(* Logix 5000 project; controller PLC_MCC1300_75F1 vendor 1 type 14 code 166 rev 32.11; software revision 32.04; part 40 of 83 *)
(* tags used below, declared in another part *)
   CONST_rgdDestMask : DINT[32];   // Destination Mask
   GP_RampSpace : GP_RampSpace;
   I : INT[128];   // Local Input Updates Input Slot 2
   TMP_d : DINT;
   TMP_dConv : DINT;
   TMP_dEndConveyorPos : DINT;
   TMP_dIndexMotor : DINT;
   TMP_dIndexNext : DINT;
   TMP_dIndexPrevious : DINT;
   TMP_dTailOnNextConveyor_cmm : DINT;
   TMP_xLastConv : BOOL;
   TMP_xOSN : DINT;
   TMP_xOSN_B : DINT;
   TMP_xOSR : DINT;
   TMP_xOSR_B : DINT;
   TMP_xSimulationActive : BOOL;
   xAlwaysOFF : BOOL;
   xAlwaysON : BOOL;
   xDebugOFF : BOOL;
   xDebugON : BOOL;
   Z300_Conveyor : UDT_StandConv[29];
   Z300_Conveyor_ALM : MAC_Conveyor_ZC_ALM[29];
   Z300_Conveyor_Conf : UDT_Conveyor_Config[29];
   Z300_Conveyor_HMW : MAC_Conveyor_ZC_HMW[29];
   Z300_Conveyor_IN_MOTION : MAC_Conveyor_ZC_IN_MOTION[29];
   Z300_LineTracking : UDT_LINE_TRACKING;
   Z301 : MAC_Zone_ML;
(* MainProgram, continued *)

ROUTINE Conv_Config   (* structured text *)
   //// CONVEYORS CONFIGURATION ////
   
   //M2CM01 (M302M1)
   Z300_Conveyor_Conf[0].dLengthConveyor_cmm := 45000;
   Z300_Conveyor_Conf[0].dWidthConveyor_cmm := 450000;
   Z300_Conveyor_Conf[0].dPitchRoller := 25000;
   Z300_Conveyor_Conf[0].dSpaceRestartPlate_cmm := 0;
   Z300_Conveyor_Conf[0].dMachineIndex := 0;
   Z300_Conveyor_Conf[0].dZoneConveyor := 1; //Z301
   Z300_Conveyor_Conf[0].dMotorNumber := 0; //Single motor
   Z300_Conveyor_Conf[0].dIndexMainSpeed := 1; //Lehr speed
   Z300_Conveyor_Conf[0].xContinuousConveyor := 1;
   Z300_Conveyor_Conf[0].xWaitGlassForStop := 0;
   Z300_Conveyor_Conf[0].rAccH_ms2 := 1.2;
   Z300_Conveyor_Conf[0].rDecH_ms2 := 1.2;
   Z300_Conveyor_Conf[0].rAccH_s := 0.75; //acceleration time with max speed 54 m/min
   Z300_Conveyor_Conf[0].rDecH_s := 0.75; //acceleration time with max speed 54 m/min
   Z300_Conveyor_Conf[0].rAccL_ms2 := 0.7;
   Z300_Conveyor_Conf[0].rDecL_ms2 := 0.7;
   Z300_Conveyor_Conf[0].rAccL_s := 1.29; //acceleration time with max speed 54 m/min
   Z300_Conveyor_Conf[0].rDecL_s := 1.29; //acceleration time with max speed 54 m/min
   Z300_Conveyor_Conf[0].xSimulationMotor := TMP_xSimulationActive;
   Z300_Conveyor_Conf[0].xLocalCleaningAllow := 0;
   Z300_Conveyor_Conf[0].xOnlyOnePlateAtTheTime := 0;
   Z300_Conveyor_Conf[0].rgxAllowedDest := CONST_rgdDestMask[0] AND CONST_rgdDestMask[1] AND CONST_rgdDestMask[2] AND CONST_rgdDestMask[3] AND CONST_rgdDestMask[4] AND CONST_rgdDestMask[5] AND CONST_rgdDestMask[6];
   Z300_Conveyor_Conf[0].rgxAllowedCullet := CONST_rgdDestMask[24];
   Z300_Conveyor_Conf[0].rgxAllowedQuality := CONST_rgdDestMask[29] AND CONST_rgdDestMask[30] AND CONST_rgdDestMask[31];
   Z300_Conveyor[0].tmOFF_DriveEnable[0].PRE := 30000;
   Z300_Conveyor[0].tmON_FeedbackTimeout[0].PRE := 2500;
   Z300_Conveyor[0].tmON_DelayReadyToMove[0].PRE := 200;
   Z300_Conveyor[0].tmON_FeedbackDriveReady[0].PRE := 1000;
   
   //M2CM02 (M302M2)
   Z300_Conveyor_Conf[1].dLengthConveyor_cmm := 31000;
   Z300_Conveyor_Conf[1].dWidthConveyor_cmm := 450000;
   Z300_Conveyor_Conf[1].dPitchRoller := 25000;
   Z300_Conveyor_Conf[1].dSpaceRestartPlate_cmm := 0;
   Z300_Conveyor_Conf[1].dMachineIndex := 1;
   Z300_Conveyor_Conf[1].dZoneConveyor := 1; //Z301
   Z300_Conveyor_Conf[1].dMotorNumber := 0; //Single motor
   Z300_Conveyor_Conf[1].dIndexMainSpeed := 1; //Lehr speed
   Z300_Conveyor_Conf[1].xContinuousConveyor := 1;
   Z300_Conveyor_Conf[1].xWaitGlassForStop := 0;
   Z300_Conveyor_Conf[1].rAccH_ms2 := 1.2;
   Z300_Conveyor_Conf[1].rDecH_ms2 := 1.2;
   Z300_Conveyor_Conf[1].rAccH_s := 0.75; //acceleration time with max speed 54 m/min
   Z300_Conveyor_Conf[1].rDecH_s := 0.75; //acceleration time with max speed 54 m/min
   Z300_Conveyor_Conf[1].rAccL_ms2 := 0.7;
   Z300_Conveyor_Conf[1].rDecL_ms2 := 0.7;
   Z300_Conveyor_Conf[1].rAccL_s := 1.29; //acceleration time with max speed 54 m/min
   Z300_Conveyor_Conf[1].rDecL_s := 1.29; //acceleration time with max speed 54 m/min
   Z300_Conveyor_Conf[1].xSimulationMotor := TMP_xSimulationActive;
   Z300_Conveyor_Conf[1].xLocalCleaningAllow := 0;
   Z300_Conveyor_Conf[1].xOnlyOnePlateAtTheTime := 0;
   Z300_Conveyor_Conf[1].rgxAllowedDest := CONST_rgdDestMask[0] AND CONST_rgdDestMask[1] AND CONST_rgdDestMask[2] AND CONST_rgdDestMask[3] AND CONST_rgdDestMask[4] AND CONST_rgdDestMask[5] AND CONST_rgdDestMask[6];
   Z300_Conveyor_Conf[1].rgxAllowedCullet := CONST_rgdDestMask[24];
   Z300_Conveyor_Conf[1].rgxAllowedQuality := CONST_rgdDestMask[29] AND CONST_rgdDestMask[30] AND CONST_rgdDestMask[31];
   Z300_Conveyor[1].tmOFF_DriveEnable[0].PRE := 30000;
   Z300_Conveyor[1].tmON_FeedbackTimeout[0].PRE := 2500;
   Z300_Conveyor[1].tmON_DelayReadyToMove[0].PRE := 200;
   Z300_Conveyor[1].tmON_FeedbackDriveReady[0].PRE := 1000;
   
   //M2CM03 (M302M3)
   Z300_Conveyor_Conf[2].dLengthConveyor_cmm := 16000;
   Z300_Conveyor_Conf[2].dWidthConveyor_cmm := 450000;
   Z300_Conveyor_Conf[2].dPitchRoller := 25000;
   Z300_Conveyor_Conf[2].dSpaceRestartPlate_cmm := 0;
   Z300_Conveyor_Conf[2].dMachineIndex := 2;
   Z300_Conveyor_Conf[2].dZoneConveyor := 1; //Z301
   Z300_Conveyor_Conf[2].dMotorNumber := 0; //Single motor
   Z300_Conveyor_Conf[2].dIndexMainSpeed := 1; //Lehr speed
   Z300_Conveyor_Conf[2].xContinuousConveyor := 1;
   Z300_Conveyor_Conf[2].xWaitGlassForStop := 0;
   Z300_Conveyor_Conf[2].rAccH_ms2 := 1.2;
   Z300_Conveyor_Conf[2].rDecH_ms2 := 1.2;
   Z300_Conveyor_Conf[2].rAccH_s := 0.75; //acceleration time with max speed 54 m/min
   Z300_Conveyor_Conf[2].rDecH_s := 0.75; //acceleration time with max speed 54 m/min
   Z300_Conveyor_Conf[2].rAccL_ms2 := 0.7;
   Z300_Conveyor_Conf[2].rDecL_ms2 := 0.7;
   Z300_Conveyor_Conf[2].rAccL_s := 1.29; //acceleration time with max speed 54 m/min
   Z300_Conveyor_Conf[2].rDecL_s := 1.29; //acceleration time with max speed 54 m/min
   Z300_Conveyor_Conf[2].xSimulationMotor := TMP_xSimulationActive;
   Z300_Conveyor_Conf[2].xLocalCleaningAllow := 0;
   Z300_Conveyor_Conf[2].xOnlyOnePlateAtTheTime := 0;
   Z300_Conveyor_Conf[2].rgxAllowedDest := CONST_rgdDestMask[0] AND CONST_rgdDestMask[1] AND CONST_rgdDestMask[2] AND CONST_rgdDestMask[3] AND CONST_rgdDestMask[4] AND CONST_rgdDestMask[5] AND CONST_rgdDestMask[6];
   Z300_Conveyor_Conf[2].rgxAllowedCullet := CONST_rgdDestMask[24];
   Z300_Conveyor_Conf[2].rgxAllowedQuality := CONST_rgdDestMask[29] AND CONST_rgdDestMask[30] AND CONST_rgdDestMask[31];
   Z300_Conveyor[2].tmOFF_DriveEnable[0].PRE := 30000;
   Z300_Conveyor[2].tmON_FeedbackTimeout[0].PRE := 2500;
   Z300_Conveyor[2].tmON_DelayReadyToMove[0].PRE := 200;
   Z300_Conveyor[2].tmON_FeedbackDriveReady[0].PRE := 1000;
   
   //M2CM04 (M302M4)
   Z300_Conveyor_Conf[3].dLengthConveyor_cmm := 47000;
   Z300_Conveyor_Conf[3].dWidthConveyor_cmm := 450000;
   Z300_Conveyor_Conf[3].dPitchRoller := 25000;
   Z300_Conveyor_Conf[3].dSpaceRestartPlate_cmm := 0;
   Z300_Conveyor_Conf[3].dMachineIndex := 3;
   Z300_Conveyor_Conf[3].dZoneConveyor := 1; //Z301
   Z300_Conveyor_Conf[3].dMotorNumber := 0; //Single motor
   Z300_Conveyor_Conf[3].dIndexMainSpeed := 1; //Lehr speed
   Z300_Conveyor_Conf[3].xContinuousConveyor := 1;
   Z300_Conveyor_Conf[3].xWaitGlassForStop := 0;
   Z300_Conveyor_Conf[3].rAccH_ms2 := 1.2;
   Z300_Conveyor_Conf[3].rDecH_ms2 := 1.2;
   Z300_Conveyor_Conf[3].rAccH_s := 0.75; //acceleration time with max speed 54 m/min
   Z300_Conveyor_Conf[3].rDecH_s := 0.75; //acceleration time with max speed 54 m/min
   Z300_Conveyor_Conf[3].rAccL_ms2 := 0.7;
   Z300_Conveyor_Conf[3].rDecL_ms2 := 0.7;
   Z300_Conveyor_Conf[3].rAccL_s := 1.29; //acceleration time with max speed 54 m/min
   Z300_Conveyor_Conf[3].rDecL_s := 1.29; //acceleration time with max speed 54 m/min
   Z300_Conveyor_Conf[3].xSimulationMotor := TMP_xSimulationActive;
   Z300_Conveyor_Conf[3].xLocalCleaningAllow := 0;
   Z300_Conveyor_Conf[3].xOnlyOnePlateAtTheTime := 0;
   Z300_Conveyor_Conf[3].rgxAllowedDest := CONST_rgdDestMask[0] AND CONST_rgdDestMask[1] AND CONST_rgdDestMask[2] AND CONST_rgdDestMask[3] AND CONST_rgdDestMask[4] AND CONST_rgdDestMask[5] AND CONST_rgdDestMask[6];
   Z300_Conveyor_Conf[3].rgxAllowedCullet := CONST_rgdDestMask[24];
   Z300_Conveyor_Conf[3].rgxAllowedQuality := CONST_rgdDestMask[29] AND CONST_rgdDestMask[30] AND CONST_rgdDestMask[31];
   Z300_Conveyor[3].tmOFF_DriveEnable[0].PRE := 30000;
   Z300_Conveyor[3].tmON_FeedbackTimeout[0].PRE := 2500;
   Z300_Conveyor[3].tmON_DelayReadyToMove[0].PRE := 200;
   Z300_Conveyor[3].tmON_FeedbackDriveReady[0].PRE := 1000;
   
   //M2CM05 (M302M5)
   Z300_Conveyor_Conf[4].dLengthConveyor_cmm := 62000;
   Z300_Conveyor_Conf[4].dWidthConveyor_cmm := 450000;
   Z300_Conveyor_Conf[4].dPitchRoller := 25000;
   Z300_Conveyor_Conf[4].dSpaceRestartPlate_cmm := 0;
   Z300_Conveyor_Conf[4].dMachineIndex := 4;
   Z300_Conveyor_Conf[4].dZoneConveyor := 1; //Z301
   Z300_Conveyor_Conf[4].dMotorNumber := 0; //Single motor
   Z300_Conveyor_Conf[4].dIndexMainSpeed := 1; //Lehr speed
   Z300_Conveyor_Conf[4].xContinuousConveyor := 1;
   Z300_Conveyor_Conf[4].xWaitGlassForStop := 0;
   Z300_Conveyor_Conf[4].rAccH_ms2 := 1.2;
   Z300_Conveyor_Conf[4].rDecH_ms2 := 1.2;
   Z300_Conveyor_Conf[4].rAccH_s := 0.75; //acceleration time with max speed 54 m/min
   Z300_Conveyor_Conf[4].rDecH_s := 0.75; //acceleration time with max speed 54 m/min
   Z300_Conveyor_Conf[4].rAccL_ms2 := 0.7;
   Z300_Conveyor_Conf[4].rDecL_ms2 := 0.7;
   Z300_Conveyor_Conf[4].rAccL_s := 1.29; //acceleration time with max speed 54 m/min
   Z300_Conveyor_Conf[4].rDecL_s := 1.29; //acceleration time with max speed 54 m/min
   Z300_Conveyor_Conf[4].xSimulationMotor := TMP_xSimulationActive;
   Z300_Conveyor_Conf[4].xLocalCleaningAllow := 0;
   Z300_Conveyor_Conf[4].xOnlyOnePlateAtTheTime := 0;
   Z300_Conveyor_Conf[4].rgxAllowedDest := CONST_rgdDestMask[0] AND CONST_rgdDestMask[1] AND CONST_rgdDestMask[2] AND CONST_rgdDestMask[3] AND CONST_rgdDestMask[4] AND CONST_rgdDestMask[5] AND CONST_rgdDestMask[6];
   Z300_Conveyor_Conf[4].rgxAllowedCullet := CONST_rgdDestMask[24];
   Z300_Conveyor_Conf[4].rgxAllowedQuality := CONST_rgdDestMask[29] AND CONST_rgdDestMask[30] AND CONST_rgdDestMask[31];
   Z300_Conveyor[4].tmOFF_DriveEnable[0].PRE := 30000;
   Z300_Conveyor[4].tmON_FeedbackTimeout[0].PRE := 2500;
   Z300_Conveyor[4].tmON_DelayReadyToMove[0].PRE := 200;
   Z300_Conveyor[4].tmON_FeedbackDriveReady[0].PRE := 1000;
   
   //M2CM06 (M302M6)
   Z300_Conveyor_Conf[5].dLengthConveyor_cmm := 93000;
   Z300_Conveyor_Conf[5].dWidthConveyor_cmm := 450000;
   Z300_Conveyor_Conf[5].dPitchRoller := 25000;
   Z300_Conveyor_Conf[5].dSpaceRestartPlate_cmm := 0;
   Z300_Conveyor_Conf[5].dMachineIndex := 5;
   Z300_Conveyor_Conf[5].dZoneConveyor := 1; //Z301
   Z300_Conveyor_Conf[5].dMotorNumber := 1; //Double motor
   Z300_Conveyor_Conf[5].dIndexMainSpeed := 3; //Special speed
   Z300_Conveyor_Conf[5].xContinuousConveyor := 1;
   Z300_Conveyor_Conf[5].xWaitGlassForStop := 0;
   Z300_Conveyor_Conf[5].rAccH_ms2 := 1.2;
   Z300_Conveyor_Conf[5].rDecH_ms2 := 1.2;
   Z300_Conveyor_Conf[5].rAccH_s := 0.75; //acceleration time with max speed 54 m/min
   Z300_Conveyor_Conf[5].rDecH_s := 0.75; //acceleration time with max speed 54 m/min
   Z300_Conveyor_Conf[5].rAccL_ms2 := 0.7;
   Z300_Conveyor_Conf[5].rDecL_ms2 := 0.7;
   Z300_Conveyor_Conf[5].rAccL_s := 1.29; //acceleration time with max speed 54 m/min
   Z300_Conveyor_Conf[5].rDecL_s := 1.29; //acceleration time with max speed 54 m/min
   Z300_Conveyor_Conf[5].xSimulationMotor := TMP_xSimulationActive;
   Z300_Conveyor_Conf[5].xLocalCleaningAllow := 0;
   Z300_Conveyor_Conf[5].xOnlyOnePlateAtTheTime := 0;
   Z300_Conveyor_Conf[5].rgxAllowedDest := CONST_rgdDestMask[0] AND CONST_rgdDestMask[1] AND CONST_rgdDestMask[2] AND CONST_rgdDestMask[3] AND CONST_rgdDestMask[4] AND CONST_rgdDestMask[5] AND CONST_rgdDestMask[6];
   Z300_Conveyor_Conf[5].rgxAllowedCullet := CONST_rgdDestMask[24];
   Z300_Conveyor_Conf[5].rgxAllowedQuality := CONST_rgdDestMask[29] AND CONST_rgdDestMask[30] AND CONST_rgdDestMask[31];
   Z300_Conveyor[5].tmOFF_DriveEnable[0].PRE := 30000;
   Z300_Conveyor[5].tmOFF_DriveEnable[1].PRE := 30000;
   Z300_Conveyor[5].tmON_FeedbackTimeout[0].PRE := 2500;
   Z300_Conveyor[5].tmON_FeedbackTimeout[1].PRE := 2500;
   Z300_Conveyor[5].tmON_DelayReadyToMove[0].PRE := 200;
   Z300_Conveyor[5].tmON_DelayReadyToMove[1].PRE := 200;
   Z300_Conveyor[5].tmON_FeedbackDriveReady[0].PRE := 1000;
   Z300_Conveyor[5].tmON_FeedbackDriveReady[1].PRE := 1000;
   
   //M2CM07 (M302M7)
   Z300_Conveyor_Conf[6].dLengthConveyor_cmm := 123000;
   Z300_Conveyor_Conf[6].dWidthConveyor_cmm := 450000;
   Z300_Conveyor_Conf[6].dPitchRoller := 25000;
   Z300_Conveyor_Conf[6].dSpaceRestartPlate_cmm := 0;
   Z300_Conveyor_Conf[6].dMachineIndex := 6;
   Z300_Conveyor_Conf[6].dZoneConveyor := 1; //Z301
   Z300_Conveyor_Conf[6].dMotorNumber := 0; //Single motor
   Z300_Conveyor_Conf[6].dIndexMainSpeed := 3; //Special speed
   Z300_Conveyor_Conf[6].xContinuousConveyor := 1;
   Z300_Conveyor_Conf[6].xWaitGlassForStop := 0;
   Z300_Conveyor_Conf[6].rAccH_ms2 := 1.2;
   Z300_Conveyor_Conf[6].rDecH_ms2 := 1.2;
   Z300_Conveyor_Conf[6].rAccH_s := 0.75; //acceleration time with max speed 54 m/min
   Z300_Conveyor_Conf[6].rDecH_s := 0.75; //acceleration time with max speed 54 m/min
   Z300_Conveyor_Conf[6].rAccL_ms2 := 0.7;
   Z300_Conveyor_Conf[6].rDecL_ms2 := 0.7;
   Z300_Conveyor_Conf[6].rAccL_s := 1.29; //acceleration time with max speed 54 m/min
   Z300_Conveyor_Conf[6].rDecL_s := 1.29; //acceleration time with max speed 54 m/min
   Z300_Conveyor_Conf[6].xSimulationMotor := TMP_xSimulationActive;
   Z300_Conveyor_Conf[6].xLocalCleaningAllow := 0;
   Z300_Conveyor_Conf[6].xOnlyOnePlateAtTheTime := 0;
   Z300_Conveyor_Conf[6].rgxAllowedDest := CONST_rgdDestMask[0] AND CONST_rgdDestMask[1] AND CONST_rgdDestMask[2] AND CONST_rgdDestMask[3] AND CONST_rgdDestMask[4] AND CONST_rgdDestMask[5] AND CONST_rgdDestMask[6];
   Z300_Conveyor_Conf[6].rgxAllowedCullet := CONST_rgdDestMask[24];
   Z300_Conveyor_Conf[6].rgxAllowedQuality := CONST_rgdDestMask[29] AND CONST_rgdDestMask[30] AND CONST_rgdDestMask[31];
   Z300_Conveyor[6].tmOFF_DriveEnable[0].PRE := 30000;
   Z300_Conveyor[6].tmON_FeedbackTimeout[0].PRE := 2500;
   Z300_Conveyor[6].tmON_DelayReadyToMove[0].PRE := 200;
   Z300_Conveyor[6].tmON_FeedbackDriveReady[0].PRE := 1000;
   
   //M2CM08 (M303M1)
   Z300_Conveyor_Conf[7].dLengthConveyor_cmm := 168000;
   Z300_Conveyor_Conf[7].dWidthConveyor_cmm := 450000;
   Z300_Conveyor_Conf[7].dPitchRoller := 25000;
   Z300_Conveyor_Conf[7].dSpaceRestartPlate_cmm := 0;
   Z300_Conveyor_Conf[7].dMachineIndex := 7;
   Z300_Conveyor_Conf[7].dZoneConveyor := 1; //Z301
   Z300_Conveyor_Conf[7].dMotorNumber := 0; //Single motor
   Z300_Conveyor_Conf[7].dIndexMainSpeed := 3; //Special speed
   Z300_Conveyor_Conf[7].xContinuousConveyor := 1;
   Z300_Conveyor_Conf[7].xWaitGlassForStop := 0;
   Z300_Conveyor_Conf[7].rAccH_ms2 := 1.2;
   Z300_Conveyor_Conf[7].rDecH_ms2 := 1.2;
   Z300_Conveyor_Conf[7].rAccH_s := 0.75; //acceleration time with max speed 54 m/min
   Z300_Conveyor_Conf[7].rDecH_s := 0.75; //acceleration time with max speed 54 m/min
   Z300_Conveyor_Conf[7].rAccL_ms2 := 0.7;
   Z300_Conveyor_Conf[7].rDecL_ms2 := 0.7;
   Z300_Conveyor_Conf[7].rAccL_s := 1.29; //acceleration time with max speed 54 m/min
   Z300_Conveyor_Conf[7].rDecL_s := 1.29; //acceleration time with max speed 54 m/min
   Z300_Conveyor_Conf[7].xSimulationMotor := TMP_xSimulationActive;
   Z300_Conveyor_Conf[7].xLocalCleaningAllow := 0;
   Z300_Conveyor_Conf[7].xOnlyOnePlateAtTheTime := 0;
   Z300_Conveyor_Conf[7].rgxAllowedDest := CONST_rgdDestMask[0] AND CONST_rgdDestMask[1] AND CONST_rgdDestMask[2] AND CONST_rgdDestMask[3] AND CONST_rgdDestMask[4] AND CONST_rgdDestMask[5] AND CONST_rgdDestMask[6];
   Z300_Conveyor_Conf[7].rgxAllowedCullet := CONST_rgdDestMask[24];
   Z300_Conveyor_Conf[7].rgxAllowedQuality := CONST_rgdDestMask[29] AND CONST_rgdDestMask[30] AND CONST_rgdDestMask[31];
   Z300_Conveyor[7].tmOFF_DriveEnable[0].PRE := 30000;
   Z300_Conveyor[7].tmON_FeedbackTimeout[0].PRE := 2500;
   Z300_Conveyor[7].tmON_DelayReadyToMove[0].PRE := 200;
   Z300_Conveyor[7].tmON_FeedbackDriveReady[0].PRE := 1000;
   
   //M2CM09 (M303M2)
   Z300_Conveyor_Conf[8].dLengthConveyor_cmm := 183000;
   Z300_Conveyor_Conf[8].dWidthConveyor_cmm := 450000;
   Z300_Conveyor_Conf[8].dPitchRoller := 25000;
   Z300_Conveyor_Conf[8].dSpaceRestartPlate_cmm := 0;
   Z300_Conveyor_Conf[8].dMachineIndex := 8;
   Z300_Conveyor_Conf[8].dZoneConveyor := 1; //Z301
   Z300_Conveyor_Conf[8].dMotorNumber := 0; //Single motor
   Z300_Conveyor_Conf[8].dIndexMainSpeed := 3; //Special speed
   Z300_Conveyor_Conf[8].xContinuousConveyor := 1;
   Z300_Conveyor_Conf[8].xWaitGlassForStop := 0;
   Z300_Conveyor_Conf[8].rAccH_ms2 := 1.2;
   Z300_Conveyor_Conf[8].rDecH_ms2 := 1.2;
   Z300_Conveyor_Conf[8].rAccH_s := 1.25; //acceleration time with max speed 90 m/min
   Z300_Conveyor_Conf[8].rDecH_s := 1.25; //acceleration time with max speed 90 m/min
   Z300_Conveyor_Conf[8].rAccL_ms2 := 0.7;
   Z300_Conveyor_Conf[8].rDecL_ms2 := 0.7;
   Z300_Conveyor_Conf[8].rAccL_s := 2.14; //acceleration time with max speed 90 m/min
   Z300_Conveyor_Conf[8].rDecL_s := 2.14; //acceleration time with max speed 90 m/min
   Z300_Conveyor_Conf[8].xSimulationMotor := TMP_xSimulationActive;
   Z300_Conveyor_Conf[8].xLocalCleaningAllow := 0;
   Z300_Conveyor_Conf[8].xOnlyOnePlateAtTheTime := 0;
   Z300_Conveyor_Conf[8].rgxAllowedDest := CONST_rgdDestMask[0] AND CONST_rgdDestMask[1] AND CONST_rgdDestMask[2] AND CONST_rgdDestMask[3] AND CONST_rgdDestMask[4] AND CONST_rgdDestMask[5] AND CONST_rgdDestMask[6];
   Z300_Conveyor_Conf[8].rgxAllowedCullet := CONST_rgdDestMask[24];
   Z300_Conveyor_Conf[8].rgxAllowedQuality := CONST_rgdDestMask[29] AND CONST_rgdDestMask[30] AND CONST_rgdDestMask[31];
   Z300_Conveyor[8].tmOFF_DriveEnable[0].PRE := 30000;
   Z300_Conveyor[8].tmON_FeedbackTimeout[0].PRE := 2500;
   Z300_Conveyor[8].tmON_DelayReadyToMove[0].PRE := 200;
   Z300_Conveyor[8].tmON_FeedbackDriveReady[0].PRE := 1000;
   
   //M2CM10 (M304M1)
   Z300_Conveyor_Conf[9].dLengthConveyor_cmm := 381000;
   Z300_Conveyor_Conf[9].dWidthConveyor_cmm := 450000;
   Z300_Conveyor_Conf[9].dPitchRoller := 25000;
   Z300_Conveyor_Conf[9].dSpaceRestartPlate_cmm := 0;
   Z300_Conveyor_Conf[9].dMachineIndex := 9;
   Z300_Conveyor_Conf[9].dZoneConveyor := 1; //Z301
   Z300_Conveyor_Conf[9].dMotorNumber := 0; //Single motor
   Z300_Conveyor_Conf[9].dIndexMainSpeed := 3; //Special speed
   Z300_Conveyor_Conf[9].xContinuousConveyor := 1;
   Z300_Conveyor_Conf[9].xWaitGlassForStop := 0;
   Z300_Conveyor_Conf[9].rAccH_ms2 := 1.2;
   Z300_Conveyor_Conf[9].rDecH_ms2 := 1.2;
   Z300_Conveyor_Conf[9].rAccH_s := 1.25; //acceleration time with max speed 90 m/min
   Z300_Conveyor_Conf[9].rDecH_s := 1.25; //acceleration time with max speed 90 m/min
   Z300_Conveyor_Conf[9].rAccL_ms2 := 0.7;
   Z300_Conveyor_Conf[9].rDecL_ms2 := 0.7;
   Z300_Conveyor_Conf[9].rAccL_s := 2.14; //acceleration time with max speed 90 m/min
   Z300_Conveyor_Conf[9].rDecL_s := 2.14; //acceleration time with max speed 90 m/min
   Z300_Conveyor_Conf[9].xSimulationMotor := TMP_xSimulationActive;
   Z300_Conveyor_Conf[9].xLocalCleaningAllow := 0;
   Z300_Conveyor_Conf[9].xOnlyOnePlateAtTheTime := 0;
   Z300_Conveyor_Conf[9].rgxAllowedDest := CONST_rgdDestMask[0] AND CONST_rgdDestMask[1] AND CONST_rgdDestMask[2] AND CONST_rgdDestMask[3] AND CONST_rgdDestMask[4] AND CONST_rgdDestMask[5] AND CONST_rgdDestMask[6];
   Z300_Conveyor_Conf[9].rgxAllowedCullet := CONST_rgdDestMask[24];
   Z300_Conveyor_Conf[9].rgxAllowedQuality := CONST_rgdDestMask[29] AND CONST_rgdDestMask[30] AND CONST_rgdDestMask[31];
   Z300_Conveyor[9].tmOFF_DriveEnable[0].PRE := 30000;
   Z300_Conveyor[9].tmON_FeedbackTimeout[0].PRE := 2500;
   Z300_Conveyor[9].tmON_DelayReadyToMove[0].PRE := 200;
   Z300_Conveyor[9].tmON_FeedbackDriveReady[0].PRE := 1000;
   
   //M2CM11 (M305M1)
   Z300_Conveyor_Conf[10].dLengthConveyor_cmm := 381000;
   Z300_Conveyor_Conf[10].dWidthConveyor_cmm := 450000;
   Z300_Conveyor_Conf[10].dPitchRoller := 25000;
   Z300_Conveyor_Conf[10].dSpaceRestartPlate_cmm := 0;
   Z300_Conveyor_Conf[10].dMachineIndex := 10;
   Z300_Conveyor_Conf[10].dZoneConveyor := 1; //Z301
   Z300_Conveyor_Conf[10].dMotorNumber := 0; //Single motor
   Z300_Conveyor_Conf[10].dIndexMainSpeed := 3; //Special speed
   Z300_Conveyor_Conf[10].xContinuousConveyor := 1;
   Z300_Conveyor_Conf[10].xWaitGlassForStop := 0;
   Z300_Conveyor_Conf[10].rAccH_ms2 := 1.2;
   Z300_Conveyor_Conf[10].rDecH_ms2 := 1.2;
   Z300_Conveyor_Conf[10].rAccH_s := 1.25; //acceleration time with max speed 90 m/min
   Z300_Conveyor_Conf[10].rDecH_s := 1.25; //acceleration time with max speed 90 m/min
   Z300_Conveyor_Conf[10].rAccL_ms2 := 0.7;
   Z300_Conveyor_Conf[10].rDecL_ms2 := 0.7;
   Z300_Conveyor_Conf[10].rAccL_s := 2.14; //acceleration time with max speed 90 m/min
   Z300_Conveyor_Conf[10].rDecL_s := 2.14; //acceleration time with max speed 90 m/min
   Z300_Conveyor_Conf[10].xSimulationMotor := TMP_xSimulationActive;
   Z300_Conveyor_Conf[10].xLocalCleaningAllow := 0;
   Z300_Conveyor_Conf[10].xOnlyOnePlateAtTheTime := 0;
   Z300_Conveyor_Conf[10].rgxAllowedDest := CONST_rgdDestMask[0] AND CONST_rgdDestMask[1] AND CONST_rgdDestMask[2] AND CONST_rgdDestMask[3] AND CONST_rgdDestMask[4] AND CONST_rgdDestMask[5] AND CONST_rgdDestMask[6];
   Z300_Conveyor_Conf[10].rgxAllowedCullet := CONST_rgdDestMask[24];
   Z300_Conveyor_Conf[10].rgxAllowedQuality := CONST_rgdDestMask[29] AND CONST_rgdDestMask[30] AND CONST_rgdDestMask[31];
   Z300_Conveyor[10].tmOFF_DriveEnable[0].PRE := 30000;
   Z300_Conveyor[10].tmON_FeedbackTimeout[0].PRE := 2500;
   Z300_Conveyor[10].tmON_DelayReadyToMove[0].PRE := 200;
   Z300_Conveyor[10].tmON_FeedbackDriveReady[0].PRE := 1000;
   
   //M2CM12 (M306M1)
   Z300_Conveyor_Conf[11].dLengthConveyor_cmm := 229000;
   Z300_Conveyor_Conf[11].dWidthConveyor_cmm := 450000;
   Z300_Conveyor_Conf[11].dPitchRoller := 25000;
   Z300_Conveyor_Conf[11].dSpaceRestartPlate_cmm := 0;
   Z300_Conveyor_Conf[11].dMachineIndex := 11;
   Z300_Conveyor_Conf[11].dZoneConveyor := 1; //Z301
   Z300_Conveyor_Conf[11].dMotorNumber := 1; //Double motor
   Z300_Conveyor_Conf[11].dIndexMainSpeed := 0; //Auto speed
   Z300_Conveyor_Conf[11].xContinuousConveyor := 1;
   Z300_Conveyor_Conf[11].xWaitGlassForStop := 0;
   Z300_Conveyor_Conf[11].rAccH_ms2 := 1.2;
   Z300_Conveyor_Conf[11].rDecH_ms2 := 1.2;
   Z300_Conveyor_Conf[11].rAccH_s := 1.25; //acceleration time with max speed 90 m/min
   Z300_Conveyor_Conf[11].rDecH_s := 1.25; //acceleration time with max speed 90 m/min
   Z300_Conveyor_Conf[11].rAccL_ms2 := 0.7;
   Z300_Conveyor_Conf[11].rDecL_ms2 := 0.7;
   Z300_Conveyor_Conf[11].rAccL_s := 2.14; //acceleration time with max speed 90 m/min
   Z300_Conveyor_Conf[11].rDecL_s := 2.14; //acceleration time with max speed 90 m/min
   Z300_Conveyor_Conf[11].xSimulationMotor := TMP_xSimulationActive;
   Z300_Conveyor_Conf[11].xLocalCleaningAllow := 0;
   Z300_Conveyor_Conf[11].xOnlyOnePlateAtTheTime := 0;
   Z300_Conveyor_Conf[11].rgxAllowedDest := CONST_rgdDestMask[0] AND CONST_rgdDestMask[1] AND CONST_rgdDestMask[2] AND CONST_rgdDestMask[3] AND CONST_rgdDestMask[4] AND CONST_rgdDestMask[5] AND CONST_rgdDestMask[6];
   Z300_Conveyor_Conf[11].rgxAllowedCullet := CONST_rgdDestMask[24];
   Z300_Conveyor_Conf[11].rgxAllowedQuality := CONST_rgdDestMask[29] AND CONST_rgdDestMask[30] AND CONST_rgdDestMask[31];
   Z300_Conveyor[11].tmOFF_DriveEnable[0].PRE := 30000;
   Z300_Conveyor[11].tmOFF_DriveEnable[1].PRE := 30000;
   Z300_Conveyor[11].tmON_FeedbackTimeout[0].PRE := 2500;
   Z300_Conveyor[11].tmON_FeedbackTimeout[1].PRE := 2500;
   Z300_Conveyor[11].tmON_DelayReadyToMove[0].PRE := 200;
   Z300_Conveyor[11].tmON_DelayReadyToMove[1].PRE := 200;
   Z300_Conveyor[11].tmON_FeedbackDriveReady[0].PRE := 1000;
   Z300_Conveyor[11].tmON_FeedbackDriveReady[1].PRE := 1000;
   
   //M307AM1
   Z300_Conveyor_Conf[12].dLengthConveyor_cmm := 58000;
   Z300_Conveyor_Conf[12].dWidthConveyor_cmm := 450000;
   Z300_Conveyor_Conf[12].dPitchRoller := 25000;
   Z300_Conveyor_Conf[12].dSpaceRestartPlate_cmm := 0;
   Z300_Conveyor_Conf[12].dMachineIndex := 12;
   Z300_Conveyor_Conf[12].dZoneConveyor := 1; //Z301
   Z300_Conveyor_Conf[12].dMotorNumber := 0; //Single motor
   Z300_Conveyor_Conf[12].dIndexMainSpeed := 0; //Auto speed
   Z300_Conveyor_Conf[12].xContinuousConveyor := 1;
   Z300_Conveyor_Conf[12].xWaitGlassForStop := 0;
   Z300_Conveyor_Conf[12].rAccH_ms2 := 1.2;
   Z300_Conveyor_Conf[12].rDecH_ms2 := 1.2;
   Z300_Conveyor_Conf[12].rAccH_s := 1.25; //acceleration time with max speed 90 m/min
   Z300_Conveyor_Conf[12].rDecH_s := 1.25; //acceleration time with max speed 90 m/min
   Z300_Conveyor_Conf[12].rAccL_ms2 := 0.7;
   Z300_Conveyor_Conf[12].rDecL_ms2 := 0.7;
   Z300_Conveyor_Conf[12].rAccL_s := 2.14; //acceleration time with max speed 90 m/min
   Z300_Conveyor_Conf[12].rDecL_s := 2.14; //acceleration time with max speed 90 m/min
   Z300_Conveyor_Conf[12].xSimulationMotor := TMP_xSimulationActive;
   Z300_Conveyor_Conf[12].xLocalCleaningAllow := 0;
   Z300_Conveyor_Conf[12].xOnlyOnePlateAtTheTime := 0;
   Z300_Conveyor_Conf[12].rgxAllowedDest := CONST_rgdDestMask[0] AND CONST_rgdDestMask[1] AND CONST_rgdDestMask[2] AND CONST_rgdDestMask[3] AND CONST_rgdDestMask[4] AND CONST_rgdDestMask[5] AND CONST_rgdDestMask[6];
   Z300_Conveyor_Conf[12].rgxAllowedCullet := CONST_rgdDestMask[24];
   Z300_Conveyor_Conf[12].rgxAllowedQuality := CONST_rgdDestMask[29] AND CONST_rgdDestMask[30] AND CONST_rgdDestMask[31];
   Z300_Conveyor[12].tmOFF_DriveEnable[0].PRE := 30000;
   Z300_Conveyor[12].tmON_FeedbackTimeout[0].PRE := 2500;
   Z300_Conveyor[12].tmON_DelayReadyToMove[0].PRE := 200;
   Z300_Conveyor[12].tmON_FeedbackDriveReady[0].PRE := 1000;
   
   //M307AM2
   Z300_Conveyor_Conf[13].dLengthConveyor_cmm := 60000;
   Z300_Conveyor_Conf[13].dWidthConveyor_cmm := 450000;
   Z300_Conveyor_Conf[13].dPitchRoller := 25000;
   Z300_Conveyor_Conf[13].dSpaceRestartPlate_cmm := 0;
   Z300_Conveyor_Conf[13].dMachineIndex := 13;
   Z300_Conveyor_Conf[13].dZoneConveyor := 1; //Z301
   Z300_Conveyor_Conf[13].dMotorNumber := 1; //Double motor
   Z300_Conveyor_Conf[13].dIndexMainSpeed := 0; //Auto speed
   Z300_Conveyor_Conf[13].xContinuousConveyor := 1;
   Z300_Conveyor_Conf[13].xWaitGlassForStop := 0;
   Z300_Conveyor_Conf[13].rAccH_ms2 := 1.2;
   Z300_Conveyor_Conf[13].rDecH_ms2 := 1.2;
   Z300_Conveyor_Conf[13].rAccH_s := 1.25; //acceleration time with max speed 90 m/min
   Z300_Conveyor_Conf[13].rDecH_s := 1.25; //acceleration time with max speed 90 m/min
   Z300_Conveyor_Conf[13].rAccL_ms2 := 0.7;
   Z300_Conveyor_Conf[13].rDecL_ms2 := 0.7;
   Z300_Conveyor_Conf[13].rAccL_s := 2.14; //acceleration time with max speed 90 m/min
   Z300_Conveyor_Conf[13].rDecL_s := 2.14; //acceleration time with max speed 90 m/min
   Z300_Conveyor_Conf[13].xSimulationMotor := TMP_xSimulationActive;
   Z300_Conveyor_Conf[13].xLocalCleaningAllow := 0;
   Z300_Conveyor_Conf[13].xOnlyOnePlateAtTheTime := 0;
   Z300_Conveyor_Conf[13].rgxAllowedDest := CONST_rgdDestMask[0] AND CONST_rgdDestMask[1] AND CONST_rgdDestMask[2] AND CONST_rgdDestMask[3] AND CONST_rgdDestMask[4] AND CONST_rgdDestMask[5] AND CONST_rgdDestMask[6];
   Z300_Conveyor_Conf[13].rgxAllowedCullet := CONST_rgdDestMask[24];
   Z300_Conveyor_Conf[13].rgxAllowedQuality := CONST_rgdDestMask[29] AND CONST_rgdDestMask[30] AND CONST_rgdDestMask[31];
   Z300_Conveyor[13].tmOFF_DriveEnable[0].PRE := 30000;
   Z300_Conveyor[13].tmOFF_DriveEnable[1].PRE := 30000;
   Z300_Conveyor[13].tmON_FeedbackTimeout[0].PRE := 2500;
   Z300_Conveyor[13].tmON_FeedbackTimeout[1].PRE := 2500;
   Z300_Conveyor[13].tmON_DelayReadyToMove[0].PRE := 200;
   Z300_Conveyor[13].tmON_DelayReadyToMove[1].PRE := 200;
   Z300_Conveyor[13].tmON_FeedbackDriveReady[0].PRE := 1000;
   Z300_Conveyor[13].tmON_FeedbackDriveReady[1].PRE := 1000;
   
   //M307AM3
   Z300_Conveyor_Conf[14].dLengthConveyor_cmm := 90000;
   Z300_Conveyor_Conf[14].dWidthConveyor_cmm := 450000;
   Z300_Conveyor_Conf[14].dPitchRoller := 25000;
   Z300_Conveyor_Conf[14].dSpaceRestartPlate_cmm := 0;
   Z300_Conveyor_Conf[14].dMachineIndex := 14;
   Z300_Conveyor_Conf[14].dZoneConveyor := 1; //Z301
   Z300_Conveyor_Conf[14].dMotorNumber := 1; //Double motor
   Z300_Conveyor_Conf[14].dIndexMainSpeed := 0; //Auto speed
   Z300_Conveyor_Conf[14].xContinuousConveyor := 1;
   Z300_Conveyor_Conf[14].xWaitGlassForStop := 0;
   Z300_Conveyor_Conf[14].rAccH_ms2 := 1.2;
   Z300_Conveyor_Conf[14].rDecH_ms2 := 1.2;
   Z300_Conveyor_Conf[14].rAccH_s := 1.25; //acceleration time with max speed 90 m/min
   Z300_Conveyor_Conf[14].rDecH_s := 1.25; //acceleration time with max speed 90 m/min
   Z300_Conveyor_Conf[14].rAccL_ms2 := 0.7;
   Z300_Conveyor_Conf[14].rDecL_ms2 := 0.7;
   Z300_Conveyor_Conf[14].rAccL_s := 2.14; //acceleration time with max speed 90 m/min
   Z300_Conveyor_Conf[14].rDecL_s := 2.14; //acceleration time with max speed 90 m/min
   Z300_Conveyor_Conf[14].xSimulationMotor := TMP_xSimulationActive;
   Z300_Conveyor_Conf[14].xLocalCleaningAllow := 0;
   Z300_Conveyor_Conf[14].xOnlyOnePlateAtTheTime := 0;
   Z300_Conveyor_Conf[14].rgxAllowedDest := CONST_rgdDestMask[0] AND CONST_rgdDestMask[1] AND CONST_rgdDestMask[2] AND CONST_rgdDestMask[3] AND CONST_rgdDestMask[4] AND CONST_rgdDestMask[5] AND CONST_rgdDestMask[6];
   Z300_Conveyor_Conf[14].rgxAllowedCullet := CONST_rgdDestMask[24];
   Z300_Conveyor_Conf[14].rgxAllowedQuality := CONST_rgdDestMask[29] AND CONST_rgdDestMask[30] AND CONST_rgdDestMask[31];
   Z300_Conveyor[14].tmOFF_DriveEnable[0].PRE := 30000;
   Z300_Conveyor[14].tmOFF_DriveEnable[1].PRE := 30000;
   Z300_Conveyor[14].tmON_FeedbackTimeout[0].PRE := 2500;
   Z300_Conveyor[14].tmON_FeedbackTimeout[1].PRE := 2500;
   Z300_Conveyor[14].tmON_DelayReadyToMove[0].PRE := 200;
   Z300_Conveyor[14].tmON_DelayReadyToMove[1].PRE := 200;
   Z300_Conveyor[14].tmON_FeedbackDriveReady[0].PRE := 1000;
   Z300_Conveyor[14].tmON_FeedbackDriveReady[1].PRE := 1000;
   
   //M307AM4
   Z300_Conveyor_Conf[15].dLengthConveyor_cmm := 150000;
   Z300_Conveyor_Conf[15].dWidthConveyor_cmm := 450000;
   Z300_Conveyor_Conf[15].dPitchRoller := 25000;
   Z300_Conveyor_Conf[15].dSpaceRestartPlate_cmm := 0;
   Z300_Conveyor_Conf[15].dMachineIndex := 15;
   Z300_Conveyor_Conf[15].dZoneConveyor := 1; //Z301
   Z300_Conveyor_Conf[15].dMotorNumber := 0; //Single motor
   Z300_Conveyor_Conf[15].dIndexMainSpeed := 0; //Auto speed
   Z300_Conveyor_Conf[15].xContinuousConveyor := 1;
   Z300_Conveyor_Conf[15].xWaitGlassForStop := 0;
   Z300_Conveyor_Conf[15].rAccH_ms2 := 1.2;
   Z300_Conveyor_Conf[15].rDecH_ms2 := 1.2;
   Z300_Conveyor_Conf[15].rAccH_s := 1.25; //acceleration time with max speed 90 m/min
   Z300_Conveyor_Conf[15].rDecH_s := 1.25; //acceleration time with max speed 90 m/min
   Z300_Conveyor_Conf[15].rAccL_ms2 := 0.7;
   Z300_Conveyor_Conf[15].rDecL_ms2 := 0.7;
   Z300_Conveyor_Conf[15].rAccL_s := 2.14; //acceleration time with max speed 90 m/min
   Z300_Conveyor_Conf[15].rDecL_s := 2.14; //acceleration time with max speed 90 m/min
   Z300_Conveyor_Conf[15].xSimulationMotor := TMP_xSimulationActive;
   Z300_Conveyor_Conf[15].xLocalCleaningAllow := 0;
   Z300_Conveyor_Conf[15].xOnlyOnePlateAtTheTime := 0;
   Z300_Conveyor_Conf[15].rgxAllowedDest := CONST_rgdDestMask[0] AND CONST_rgdDestMask[1] AND CONST_rgdDestMask[2] AND CONST_rgdDestMask[3] AND CONST_rgdDestMask[4] AND CONST_rgdDestMask[5] AND CONST_rgdDestMask[6];
   Z300_Conveyor_Conf[15].rgxAllowedCullet := CONST_rgdDestMask[24];
   Z300_Conveyor_Conf[15].rgxAllowedQuality := CONST_rgdDestMask[29] AND CONST_rgdDestMask[30] AND CONST_rgdDestMask[31];
   Z300_Conveyor[15].tmOFF_DriveEnable[0].PRE := 30000;
   Z300_Conveyor[15].tmON_FeedbackTimeout[0].PRE := 2500;
   Z300_Conveyor[15].tmON_DelayReadyToMove[0].PRE := 200;
   Z300_Conveyor[15].tmON_FeedbackDriveReady[0].PRE := 1000;
   
   //M307BM1
   Z300_Conveyor_Conf[16].dLengthConveyor_cmm := 238000;
   Z300_Conveyor_Conf[16].dWidthConveyor_cmm := 450000;
   Z300_Conveyor_Conf[16].dPitchRoller := 25000;
   Z300_Conveyor_Conf[16].dSpaceRestartPlate_cmm := 0;
   Z300_Conveyor_Conf[16].dMachineIndex := 16;
   Z300_Conveyor_Conf[16].dZoneConveyor := 1; //Z301
   Z300_Conveyor_Conf[16].dMotorNumber := 0; //Single motor
   Z300_Conveyor_Conf[16].dIndexMainSpeed := 0; //Auto speed
   Z300_Conveyor_Conf[16].xContinuousConveyor := 1;
   Z300_Conveyor_Conf[16].xWaitGlassForStop := 0;
   Z300_Conveyor_Conf[16].rAccH_ms2 := 1.2;
   Z300_Conveyor_Conf[16].rDecH_ms2 := 1.2;
   Z300_Conveyor_Conf[16].rAccH_s := 1.25; //acceleration time with max speed 90 m/min
   Z300_Conveyor_Conf[16].rDecH_s := 1.25; //acceleration time with max speed 90 m/min
   Z300_Conveyor_Conf[16].rAccL_ms2 := 0.7;
   Z300_Conveyor_Conf[16].rDecL_ms2 := 0.7;
   Z300_Conveyor_Conf[16].rAccL_s := 2.14; //acceleration time with max speed 90 m/min
   Z300_Conveyor_Conf[16].rDecL_s := 2.14; //acceleration time with max speed 90 m/min
   Z300_Conveyor_Conf[16].xSimulationMotor := TMP_xSimulationActive;
   Z300_Conveyor_Conf[16].xLocalCleaningAllow := 0;
   Z300_Conveyor_Conf[16].xOnlyOnePlateAtTheTime := 0;
   Z300_Conveyor_Conf[16].rgxAllowedDest := CONST_rgdDestMask[0] AND CONST_rgdDestMask[1] AND CONST_rgdDestMask[2] AND CONST_rgdDestMask[3];
   Z300_Conveyor_Conf[16].rgxAllowedCullet := CONST_rgdDestMask[24];
   Z300_Conveyor_Conf[16].rgxAllowedQuality := CONST_rgdDestMask[29] AND CONST_rgdDestMask[30] AND CONST_rgdDestMask[31];
   Z300_Conveyor[16].tmOFF_DriveEnable[0].PRE := 30000;
   Z300_Conveyor[16].tmON_FeedbackTimeout[0].PRE := 2500;
   Z300_Conveyor[16].tmON_DelayReadyToMove[0].PRE := 200;
   Z300_Conveyor[16].tmON_FeedbackDriveReady[0].PRE := 1000;
   
   //M307CM1
   Z300_Conveyor_Conf[17].dLengthConveyor_cmm := 238000;
   Z300_Conveyor_Conf[17].dWidthConveyor_cmm := 450000;
   Z300_Conveyor_Conf[17].dPitchRoller := 25000;
   Z300_Conveyor_Conf[17].dSpaceRestartPlate_cmm := 0;
   Z300_Conveyor_Conf[17].dMachineIndex := 17;
   Z300_Conveyor_Conf[17].dZoneConveyor := 1; //Z301
   Z300_Conveyor_Conf[17].dMotorNumber := 0; //Single motor
   Z300_Conveyor_Conf[17].dIndexMainSpeed := 0; //Auto speed
   Z300_Conveyor_Conf[17].xContinuousConveyor := 1;
   Z300_Conveyor_Conf[17].xWaitGlassForStop := 0;
   Z300_Conveyor_Conf[17].rAccH_ms2 := 1.2;
   Z300_Conveyor_Conf[17].rDecH_ms2 := 1.2;
   Z300_Conveyor_Conf[17].rAccH_s := 1.25; //acceleration time with max speed 90 m/min
   Z300_Conveyor_Conf[17].rDecH_s := 1.25; //acceleration time with max speed 90 m/min
   Z300_Conveyor_Conf[17].rAccL_ms2 := 0.7;
   Z300_Conveyor_Conf[17].rDecL_ms2 := 0.7;
   Z300_Conveyor_Conf[17].rAccL_s := 2.14; //acceleration time with max speed 90 m/min
   Z300_Conveyor_Conf[17].rDecL_s := 2.14; //acceleration time with max speed 90 m/min
   Z300_Conveyor_Conf[17].xSimulationMotor := TMP_xSimulationActive;
   Z300_Conveyor_Conf[17].xLocalCleaningAllow := 0;
   Z300_Conveyor_Conf[17].xOnlyOnePlateAtTheTime := 0;
   Z300_Conveyor_Conf[17].rgxAllowedDest := CONST_rgdDestMask[0] AND CONST_rgdDestMask[1] AND CONST_rgdDestMask[2] AND CONST_rgdDestMask[3] AND CONST_rgdDestMask[4] AND CONST_rgdDestMask[5] AND CONST_rgdDestMask[6];
   Z300_Conveyor_Conf[17].rgxAllowedCullet := CONST_rgdDestMask[24];
   Z300_Conveyor_Conf[17].rgxAllowedQuality := CONST_rgdDestMask[29] AND CONST_rgdDestMask[30] AND CONST_rgdDestMask[31];
   Z300_Conveyor[17].tmOFF_DriveEnable[0].PRE := 30000;
   Z300_Conveyor[17].tmON_FeedbackTimeout[0].PRE := 2500;
   Z300_Conveyor[17].tmON_DelayReadyToMove[0].PRE := 200;
   Z300_Conveyor[17].tmON_FeedbackDriveReady[0].PRE := 1000;
   
   ////END OF CONTINUOUS ZONE
   
   //M307DM1
   Z300_Conveyor_Conf[18].dLengthConveyor_cmm := 238000;
   Z300_Conveyor_Conf[18].dWidthConveyor_cmm := 450000;
   Z300_Conveyor_Conf[18].dPitchRoller := 25000;
   Z300_Conveyor_Conf[18].dSpaceRestartPlate_cmm := 200000;
   Z300_Conveyor_Conf[18].dMachineIndex := 18;
   Z300_Conveyor_Conf[18].dZoneConveyor := 1; //Z301
   Z300_Conveyor_Conf[18].dMotorNumber := 1; //Double motor
   Z300_Conveyor_Conf[18].dIndexMainSpeed := 0; //Auto speed
   Z300_Conveyor_Conf[18].xContinuousConveyor := 0;
   Z300_Conveyor_Conf[18].xWaitGlassForStop := 1;
   Z300_Conveyor_Conf[18].rAccH_ms2 := 1.2;
   Z300_Conveyor_Conf[18].rDecH_ms2 := 1.2;
   Z300_Conveyor_Conf[18].rAccH_s := 1.25; //acceleration time with max speed 90 m/min
   Z300_Conveyor_Conf[18].rDecH_s := 1.25; //acceleration time with max speed 90 m/min
   Z300_Conveyor_Conf[18].rAccL_ms2 := 0.7;
   Z300_Conveyor_Conf[18].rDecL_ms2 := 0.7;
   Z300_Conveyor_Conf[18].rAccL_s := 2.14; //acceleration time with max speed 90 m/min
   Z300_Conveyor_Conf[18].rDecL_s := 2.14; //acceleration time with max speed 90 m/min
   Z300_Conveyor_Conf[18].xSimulationMotor := TMP_xSimulationActive;
   Z300_Conveyor_Conf[18].xLocalCleaningAllow := 0;
   Z300_Conveyor_Conf[18].xOnlyOnePlateAtTheTime := 0;
   Z300_Conveyor_Conf[18].rgxAllowedDest := CONST_rgdDestMask[0] AND CONST_rgdDestMask[1] AND CONST_rgdDestMask[2] AND CONST_rgdDestMask[3] AND CONST_rgdDestMask[4] AND CONST_rgdDestMask[5] AND CONST_rgdDestMask[6];
   Z300_Conveyor_Conf[18].rgxAllowedCullet := CONST_rgdDestMask[24];
   Z300_Conveyor_Conf[18].rgxAllowedQuality := CONST_rgdDestMask[29] AND CONST_rgdDestMask[30] AND CONST_rgdDestMask[31];
   Z300_Conveyor[18].tmOFF_DriveEnable[0].PRE := 30000;
   Z300_Conveyor[18].tmOFF_DriveEnable[1].PRE := 30000;
   Z300_Conveyor[18].tmON_FeedbackTimeout[0].PRE := 2500;
   Z300_Conveyor[18].tmON_FeedbackTimeout[1].PRE := 2500;
   Z300_Conveyor[18].tmON_DelayReadyToMove[0].PRE := 200;
   Z300_Conveyor[18].tmON_DelayReadyToMove[1].PRE := 200;
   Z300_Conveyor[18].tmON_FeedbackDriveReady[0].PRE := 1000;
   Z300_Conveyor[18].tmON_FeedbackDriveReady[1].PRE := 1000;